REGION Network 5: PODAJANJE PLOŠČICE
   RUNG wire#powerrail
      Contact( #JeVRočnemNačinu )
      { S7_Templates := "SrcType := Int" } EQ_Contact(in1 := #stCilindra, in2 := 5)
      wire#w1
      Contact( #"TIPPEN_-" )
      S_Coil( #"Y1/2" )
      R_Coil( #"Y1/2_2" )
   END_RUNG
   RUNG wire#w1
      Contact( #"TIPPEN_+" )
      Contact( "FB_KEYENCE_GT2_ODMIKVARJENJA".oPoz1Dosezena )
      Contact( "FB_KEYENCE_GT2_ODMIKVARJENJA".oPoz1Dosezena )
      Contact( "Y1/4_odmičniCilinderVarjenje_GOR" )
      R_Coil( #"Y1/2" )
      S_Coil( #"Y1/2_2" )
   END_RUNG
   // the same network as SCL:
   #_w1 := #JeVRočnemNačinu AND (#stCilindra = 5);
   IF #_w1 AND #"TIPPEN_-" THEN
       #"Y1/2" := TRUE;
       #"Y1/2_2" := FALSE;
   END_IF;
   IF #_w1 AND #"TIPPEN_+" AND "FB_KEYENCE_GT2_ODMIKVARJENJA".oPoz1Dosezena AND "FB_KEYENCE_GT2_ODMIKVARJENJA".oPoz1Dosezena AND "Y1/4_odmičniCilinderVarjenje_GOR" THEN
       #"Y1/2" := FALSE;
       #"Y1/2_2" := TRUE;
   END_IF;
END_REGION

REGION Network 6: DVIG/SPUST ELEKTRODE
   RUNG wire#powerrail
      Contact( #JeVRočnemNačinu )
      { S7_Templates := "SrcType := Int" } EQ_Contact(in1 := #stCilindra, in2 := 6)
      wire#w1
      Contact( #"TIPPEN_-" )
      S_Coil( #"Y1/4_1" )
      R_Coil( #"Y1/4_2" )
   END_RUNG
   RUNG wire#w1
      Contact( #"TIPPEN_+" )
      R_Coil( #"Y1/4_1" )
      S_Coil( #"Y1/4_2" )
   END_RUNG
   // the same network as SCL:
   #_w1 := #JeVRočnemNačinu AND (#stCilindra = 6);
   IF #_w1 AND #"TIPPEN_-" THEN
       #"Y1/4_1" := TRUE;
       #"Y1/4_2" := FALSE;
   END_IF;
   IF #_w1 AND #"TIPPEN_+" THEN
       #"Y1/4_1" := FALSE;
       #"Y1/4_2" := TRUE;
   END_IF;
END_REGION

REGION Network 7: PORAVNAVA KONTAKTA
   RUNG wire#powerrail
      Contact( #JeVRočnemNačinu )
      { S7_Templates := "SrcType := Int" } EQ_Contact(in1 := #stCilindra, in2 := 7)
      wire#w1
      Contact( #"TIPPEN_-" )
      S_Coil( #"Y2/3_2" )
      R_Coil( #"Y2/3_1" )
   END_RUNG
   RUNG wire#w1
      Contact( #"TIPPEN_+" )
      R_Coil( #"Y2/3_2" )
      S_Coil( #"Y2/3_1" )
   END_RUNG
   // the same network as SCL:
   #_w1 := #JeVRočnemNačinu AND (#stCilindra = 7);
   IF #_w1 AND #"TIPPEN_-" THEN
       #"Y2/3_2" := TRUE;
       #"Y2/3_1" := FALSE;
   END_IF;
   IF #_w1 AND #"TIPPEN_+" THEN
       #"Y2/3_2" := FALSE;
       #"Y2/3_1" := TRUE;
   END_IF;
END_REGION

REGION Network 8: ODKLEP/ZAKLEP KONUSA - ROTACISKA MIZA
   RUNG wire#powerrail
      Contact( #JeVRočnemNačinu )
      { S7_Templates := "SrcType := Int" } EQ_Contact(in1 := #stCilindra, in2 := 8)
      wire#w1
      Contact( #"TIPPEN_-" )
      R_Coil( #"Y3/1_1" )
   END_RUNG
   RUNG wire#w1
      Contact( #"TIPPEN_+" )
      S_Coil( #"Y3/1_1" )
   END_RUNG
   // the same network as SCL:
   #_w1 := #JeVRočnemNačinu AND (#stCilindra = 8);
   IF #_w1 AND #"TIPPEN_-" THEN #"Y3/1_1" := FALSE; END_IF;
   IF #_w1 AND #"TIPPEN_+" THEN #"Y3/1_1" := TRUE; END_IF;
END_REGION

REGION Network 9: ODKLEP/ZAKLEP VSTAVLJANJA KOMADA V MIZO - ODKLEP ZA VSTAVLJANJE
   RUNG wire#powerrail
      Contact( #JeVRočnemNačinu )
      { S7_Templates := "SrcType := Int" } EQ_Contact(in1 := #stCilindra, in2 := 9)
      wire#w1
      Contact( #"TIPPEN_-" )
      R_Coil( #"Y3/3_1" )
   END_RUNG
   RUNG wire#w1
      Contact( #"TIPPEN_+" )
      S_Coil( #"Y3/3_1" )
   END_RUNG
   // the same network as SCL:
   #_w1 := #JeVRočnemNačinu AND (#stCilindra = 9);
   IF #_w1 AND #"TIPPEN_-" THEN #"Y3/3_1" := FALSE; END_IF;
   IF #_w1 AND #"TIPPEN_+" THEN #"Y3/3_1" := TRUE; END_IF;
END_REGION

REGION Network 10: ODKLEP/ZAKLEP DRŽALA IZMETA KOMADA
   RUNG wire#powerrail
      Contact( #JeVRočnemNačinu )
      { S7_Templates := "SrcType := Int" } EQ_Contact(in1 := #stCilindra, in2 := 10)
      wire#w1
      Contact( #"TIPPEN_-" )
      R_Coil( #"Y4/3_1" )
   END_RUNG
   RUNG wire#w1
      Contact( #"TIPPEN_+" )
      S_Coil( #"Y4/3_1" )
   END_RUNG
   // the same network as SCL:
   #_w1 := #JeVRočnemNačinu AND (#stCilindra = 10);
   IF #_w1 AND #"TIPPEN_-" THEN #"Y4/3_1" := FALSE; END_IF;
   IF #_w1 AND #"TIPPEN_+" THEN #"Y4/3_1" := TRUE; END_IF;
END_REGION

REGION Network 11: IZMET KOMADA
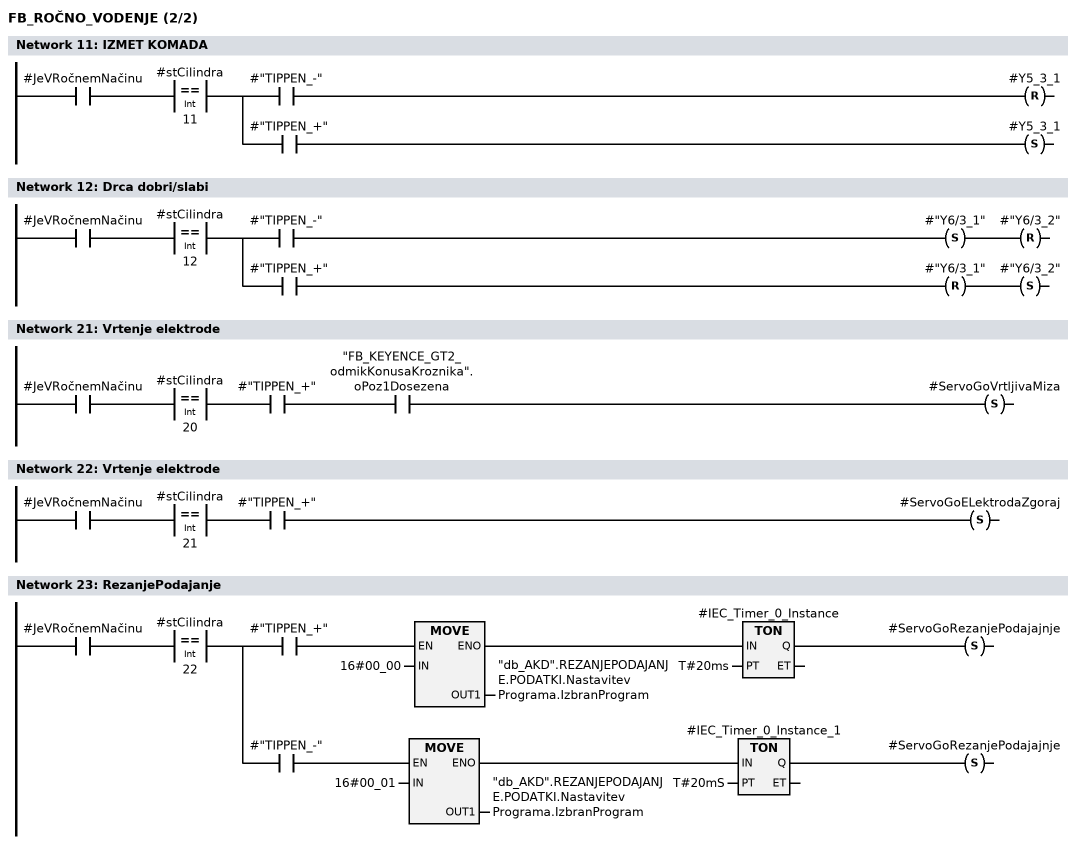
   RUNG wire#powerrail
      Contact( #JeVRočnemNačinu )
      { S7_Templates := "SrcType := Int" } EQ_Contact(in1 := #stCilindra, in2 := 11)
      wire#w1
      Contact( #"TIPPEN_-" )
      R_Coil( #Y5_3_1 )
   END_RUNG
   RUNG wire#w1
      Contact( #"TIPPEN_+" )
      S_Coil( #Y5_3_1 )
   END_RUNG
   // the same network as SCL:
   #_w1 := #JeVRočnemNačinu AND (#stCilindra = 11);
   IF #_w1 AND #"TIPPEN_-" THEN #Y5_3_1 := FALSE; END_IF;
   IF #_w1 AND #"TIPPEN_+" THEN #Y5_3_1 := TRUE; END_IF;
END_REGION

REGION Network 12: Drca dobri/slabi
   RUNG wire#powerrail
      Contact( #JeVRočnemNačinu )
      { S7_Templates := "SrcType := Int" } EQ_Contact(in1 := #stCilindra, in2 := 12)
      wire#w1
      Contact( #"TIPPEN_-" )
      S_Coil( #"Y6/3_1" )
      R_Coil( #"Y6/3_2" )
   END_RUNG
   RUNG wire#w1
      Contact( #"TIPPEN_+" )
      R_Coil( #"Y6/3_1" )
      S_Coil( #"Y6/3_2" )
   END_RUNG
   // the same network as SCL:
   #_w1 := #JeVRočnemNačinu AND (#stCilindra = 12);
   IF #_w1 AND #"TIPPEN_-" THEN
       #"Y6/3_1" := TRUE;
       #"Y6/3_2" := FALSE;
   END_IF;
   IF #_w1 AND #"TIPPEN_+" THEN
       #"Y6/3_1" := FALSE;
       #"Y6/3_2" := TRUE;
   END_IF;
END_REGION

REGION Network 21: Vrtenje elektrode
   RUNG wire#powerrail
      Contact( #JeVRočnemNačinu )
      { S7_Templates := "SrcType := Int" } EQ_Contact(in1 := #stCilindra, in2 := 20)
      Contact( #"TIPPEN_+" )
      Contact( "FB_KEYENCE_GT2_odmikKonusaKroznika".oPoz1Dosezena )
      S_Coil( #ServoGoVrtljivaMiza )
   END_RUNG
   // the same network as SCL:
   IF #JeVRočnemNačinu AND (#stCilindra = 20) AND #"TIPPEN_+" AND "FB_KEYENCE_GT2_odmikKonusaKroznika".oPoz1Dosezena THEN
       #ServoGoVrtljivaMiza := TRUE;
   END_IF;
END_REGION

REGION Network 22: Vrtenje elektrode
   RUNG wire#powerrail
      Contact( #JeVRočnemNačinu )
      { S7_Templates := "SrcType := Int" } EQ_Contact(in1 := #stCilindra, in2 := 21)
      Contact( #"TIPPEN_+" )
      S_Coil( #ServoGoELektrodaZgoraj )
   END_RUNG
   // the same network as SCL:
   IF #JeVRočnemNačinu AND (#stCilindra = 21) AND #"TIPPEN_+" THEN #ServoGoELektrodaZgoraj := TRUE; END_IF;
END_REGION

REGION Network 23: RezanjePodajanje
   #_w1 := #JeVRočnemNačinu AND (#stCilindra = 22);
   #_w2 := #_w1 AND #"TIPPEN_+";
   IF #_w2 THEN "db_AKD".REZANJEPODAJANJE.PODATKI.NastavitevPrograma.IzbranProgram := 16#00_00; END_IF;
   #IEC_Timer_0_Instance(IN := #_w2, PT := T#20ms);   // TON
   IF #IEC_Timer_0_Instance.Q THEN #ServoGoRezanjePodajajnje := TRUE; END_IF;
   #_w3 := #_w1 AND #"TIPPEN_-";
   IF #_w3 THEN "db_AKD".REZANJEPODAJANJE.PODATKI.NastavitevPrograma.IzbranProgram := 16#00_01; END_IF;
   #IEC_Timer_0_Instance_1(IN := #_w3, PT := T#20mS);   // TON
   IF #IEC_Timer_0_Instance_1.Q THEN #ServoGoRezanjePodajajnje := TRUE; END_IF;
END_REGION
END_FUNCTION_BLOCK

FUNCTION_BLOCK "FB_KEYENCE_GT2"   // FB12, LAD
{ S7_Optimized_Access := 'TRUE' }
VERSION : 0.1
   VAR_INPUT
      w_inAddr : DWord;   // VALUE| VALUE|VALUE|BDC1-4
      iPoz1 : DInt;
      iPoz2 : DInt;
      iPoz4 : DInt;
      iPoz3 : DInt;
      HISTEREZA : Int := 800;
      tol1 : Int;
      tol2 : Int;
      tol3 : Int;
      tol4 : Int;
   END_VAR
   VAR_OUTPUT
      out : UDInt;   // Rezultat int
      bBDC1 : Bool;   // Končni položaj 1
      bBDC2 : Bool;   // Končni položaj 2
      bBDC3 : Bool;   // Končni položaj 3
      bBDC4 : Bool;   // Končni položaj 4
      oPoz1Dosezena : Bool;
      oPoz2Dosezena : Bool;
      oPoz3Dosezena : Bool;
      oPoz4Dosezena : Bool;
   END_VAR
   VAR RETAIN
      w_statRor : Word;
      W_ST : Word;
   END_VAR
   VAR
      B0 : Byte;
      B1 : Byte;
   END_VAR
BEGIN

REGION Network 2 (SCL): Rezultat int
   //pozicija dosezena
   //

   #out := #w_inAddr;
   REGION POZICIJA 1
       IF (#iPoz1 - (#HISTEREZA + #tol1)) < #out AND #out < (#iPoz1 + (#HISTEREZA + #tol1)) AND #iPoz1 <> 0 THEN
           #oPoz1Dosezena := true;
   ELSE
       #oPoz1Dosezena := false;
   END_IF;
   END_REGION


   REGION POZICIJA 2
       IF (#iPoz2 - (#HISTEREZA+#tol2)) < #out AND #out < (#iPoz2 + #HISTEREZA+#tol2) AND #iPoz1 <> 0 THEN
       #oPoz2Dosezena := true;
   ELSE
       #oPoz2Dosezena := false;
   END_IF;
   END_REGION

   REGION POZICIJA 3
       IF (#iPoz3 - (#HISTEREZA+#tol3)) < #out AND #out < (#iPoz3 + #HISTEREZA+#tol3) AND #iPoz3 <> 0 THEN
           #oPoz3Dosezena := true;
       ELSE
           #oPoz3Dosezena := false;
       END_IF;
   END_REGION

   REGION POZICIJA 4
       IF (#iPoz4 - (#HISTEREZA+#tol4)) < #out AND #out < (#iPoz4 + #HISTEREZA+#tol4) AND #iPoz4 <> 0 THEN
           #oPoz4Dosezena := true;
       ELSE
           #oPoz4Dosezena := false;
       END_IF;
   END_REGION
END_REGION
END_FUNCTION_BLOCK

FUNCTION_BLOCK "FB_IZMETKOMADA"   // FB13, LAD
{ S7_Optimized_Access := 'TRUE' }
VERSION : 0.1
   VAR_OUTPUT
      VentilZaDržanjeKomada : Bool;
      VentilZaIzmetKomada : Bool;
      DržaDobriSlavi : Bool;
      DržaSlabi : Bool;
   END_VAR
   VAR_IN_OUT
      KomadiPrisotniByte : Byte;
   END_VAR
   VAR RETAIN
      statIzdelekPrisoten : Bool;
      IEC_Timer_0_Instance : TON_TIME;
      IEC_Timer_0_Instance_1 : TON_TIME;
      KoraIzmetaKoncan : Bool;
      merjerji : Array[0..10] of Bool;
   END_VAR
   VAR
      konec : Bool;
   END_VAR
BEGIN

REGION Network 2
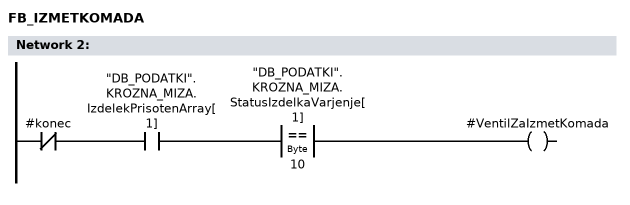
   RUNG wire#powerrail
      I_Contact( #konec )
      Contact( "DB_PODATKI".KROZNA_MIZA.IzdelekPrisotenArray[1] )
      { S7_Templates := "SrcType := Byte" } EQ_Contact(in1 := "DB_PODATKI".KROZNA_MIZA.StatusIzdelkaVarjenje[1], in2 := 10)
      Coil( #VentilZaIzmetKomada )
   END_RUNG
   // the same network as SCL:
   #VentilZaIzmetKomada := NOT #konec AND "DB_PODATKI".KROZNA_MIZA.IzdelekPrisotenArray[1] AND ("DB_PODATKI".KROZNA_MIZA.StatusIzdelkaVarjenje[1] = 10);
END_REGION
END_FUNCTION_BLOCK

FUNCTION_BLOCK "FB_VstavljanjeIzdelkaVMizo"   // FB14, LAD
{ S7_Optimized_Access := 'TRUE' }
VERSION : 0.1
   VAR_INPUT
      PogojZaVstavljanje : Bool;   // Ko na mizi ni komada
   END_VAR
   VAR_OUTPUT
      IzdelekVstavljenVMizo : Bool;
   END_VAR
   VAR RETAIN
      Korak : UInt;
   END_VAR
   VAR
      Ton : Array[0..1] of TON_TIME;
   END_VAR
   VAR_TEMP   // added for the SCL form of the ladder/FBD networks
      _w1 : Bool;
   END_VAR
BEGIN

REGION Network 1: ČajanjeZaVstavljanje
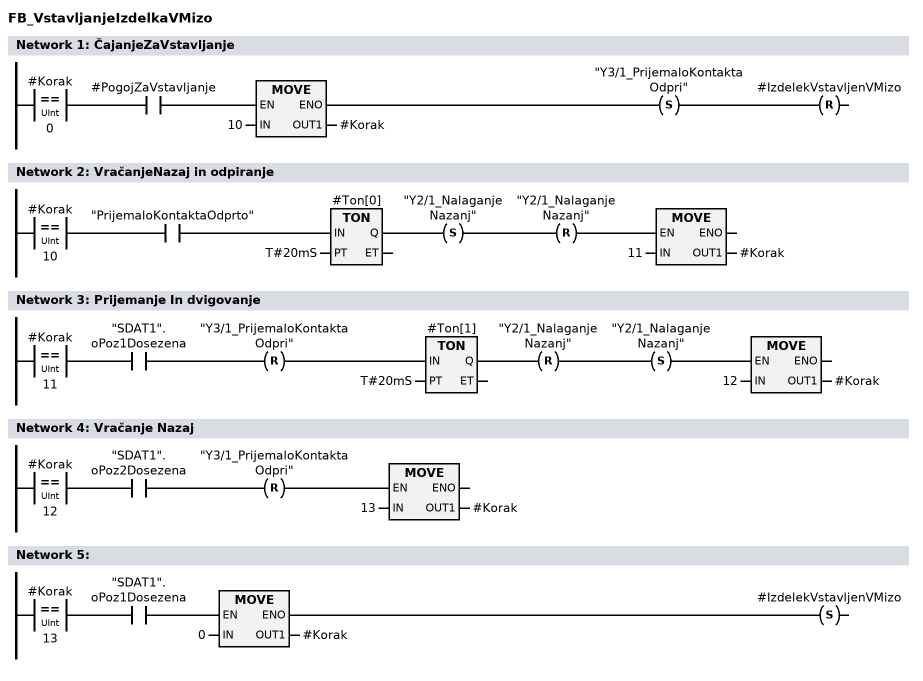
   RUNG wire#powerrail
      { S7_Templates := "SrcType := UInt" } EQ_Contact(in1 := #Korak, in2 := 0)
      Contact( #PogojZaVstavljanje )
      Move(in := 10, out1 => #Korak)
      S_Coil( "Y3/1_PrijemaloKontaktaOdpri" )
      R_Coil( #IzdelekVstavljenVMizo )
   END_RUNG
   // the same network as SCL:
   #_w1 := (#Korak = 0) AND #PogojZaVstavljanje;
   IF #_w1 THEN
       #Korak := 10;
       "Y3/1_PrijemaloKontaktaOdpri" := TRUE;
       #IzdelekVstavljenVMizo := FALSE;
   END_IF;
END_REGION

REGION Network 2: VračanjeNazaj in odpiranje
   #Ton[0].TON(IN := (#Korak = 10) AND "PrijemaloKontaktaOdprto", PT := T#20mS);
   IF #Ton[0].Q THEN
       "Y2/1_NalaganjeNazanj" := TRUE;
       "Y2/1_NalaganjeNazanj" := FALSE;
       #Korak := 11;
   END_IF;
END_REGION

REGION Network 3: Prijemanje In dvigovanje
   #_w1 := (#Korak = 11) AND "SDAT1".oPoz1Dosezena;
   IF #_w1 THEN "Y3/1_PrijemaloKontaktaOdpri" := FALSE; END_IF;
   #Ton[1].TON(IN := #_w1, PT := T#20mS);
   IF #Ton[1].Q THEN
       "Y2/1_NalaganjeNazanj" := FALSE;
       "Y2/1_NalaganjeNazanj" := TRUE;
       #Korak := 12;
   END_IF;
END_REGION

REGION Network 4: Vračanje Nazaj
   RUNG wire#powerrail
      { S7_Templates := "SrcType := UInt" } EQ_Contact(in1 := #Korak, in2 := 12)
      Contact( "SDAT1".oPoz2Dosezena )
      R_Coil( "Y3/1_PrijemaloKontaktaOdpri" )
      Move(in := 13, out1 => #Korak)
   END_RUNG
   // the same network as SCL:
   IF (#Korak = 12) AND "SDAT1".oPoz2Dosezena THEN
       "Y3/1_PrijemaloKontaktaOdpri" := FALSE;
       #Korak := 13;
   END_IF;
END_REGION

REGION Network 5
   RUNG wire#powerrail
      { S7_Templates := "SrcType := UInt" } EQ_Contact(in1 := #Korak, in2 := 13)
      Contact( "SDAT1".oPoz1Dosezena )
      Move(in := 0, out1 => #Korak)
      S_Coil( #IzdelekVstavljenVMizo )
   END_RUNG
   // the same network as SCL:
   #_w1 := (#Korak = 13) AND "SDAT1".oPoz1Dosezena;
   IF #_w1 THEN
       #Korak := 0;
       #IzdelekVstavljenVMizo := TRUE;
   END_IF;
END_REGION
END_FUNCTION_BLOCK

FUNCTION_BLOCK "FB_IOL_BANNER"   // FB15, LAD
{ S7_Optimized_Access := 'TRUE' }
VERSION : 0.1
   VAR_INPUT
      Color1 : Byte;
      ColorFlashRate : Byte;
      Color2 : Byte;
      AudioMode : Byte;
      Rotation : Bool;
      ANimationType : Byte;
      Color1Intensity : Byte;
      Color2Intensety : Byte;
   END_VAR
   VAR_OUTPUT
      oWord : DWord;
      oByte0 : Byte;
      oByte1 : Byte;
      oByte2 : Byte;
      oByte3 : Byte;
   END_VAR
   VAR
      bytes : Array[0..3] of Byte;
   END_VAR
BEGIN

REGION Network 2 (SCL)
   #bytes[0] := #Color1 + SHL(IN := #ColorFlashRate, N := 5);
   #bytes[1] := #Color2 + SHL(IN := #AudioMode, N := 5);
   #bytes[2] := #ANimationType + SHL(IN := #Color1Intensity, N := 4);
   #bytes[3] := #Color2Intensety;
   //#oWord :=#bytes[0]+SHL(IN:=#bytes[1],N:=8);
   //#oWord := ROL(IN := #oWord, N := 0);

   #oByte0 := #bytes[0];
   #oByte1 := #bytes[1];
   #oByte2 := #bytes[2];
   #oByte3 := #bytes[3];
END_REGION
END_FUNCTION_BLOCK

FUNCTION_BLOCK "FB_TekociTrak"   // FB16, LAD
{ S7_Optimized_Access := 'TRUE' }
VERSION : 0.1
   VAR_INPUT
      i_StetjeKosov : Bool;
      i_ON_OFF_TekociTrak : Bool;
      i_stevecSlabihKosov : UInt;
      i_MAX_SKATLA1 : UInt;
      i_MAX_SKATLA2 : UInt;
      i_IzprazniSKatlo1 : Bool;
      i_iprazniSkatlo2 : Bool;
   END_VAR
   VAR_OUTPUT
      o_TekočiTrak : Bool;
      o_PolnjenjeSkatle2 : Bool;
      o_Skatla1Polna : Bool;
      o_Skatla2Polna : Bool;
   END_VAR
   VAR_IN_OUT
      i_StevecSkatle1 : UInt;
      i_StevecSkatle2 : UInt;
      i_ResetNapake : Bool;
   END_VAR
   VAR RETAIN
      stat_skatla1Polna : Bool;
      stat_skatla2Polna : Bool;
      merkerji : Array[0..3] of Bool;
      IEC_Timer_0_Instance : TON_TIME;
      IEC_Timer_0_Instance_1 : TON_TIME;
      SkatliPolni : Bool;
      statPolnjenjeSkatle2 : Bool;
   END_VAR
   VAR_TEMP   // added for the SCL form of the ladder/FBD networks
      _w1 : Bool;
      _w2 : Bool;
      _w3 : Bool;
      _w4 : Bool;
   END_VAR
BEGIN

REGION Network 1: Vklop Tekocega Traka
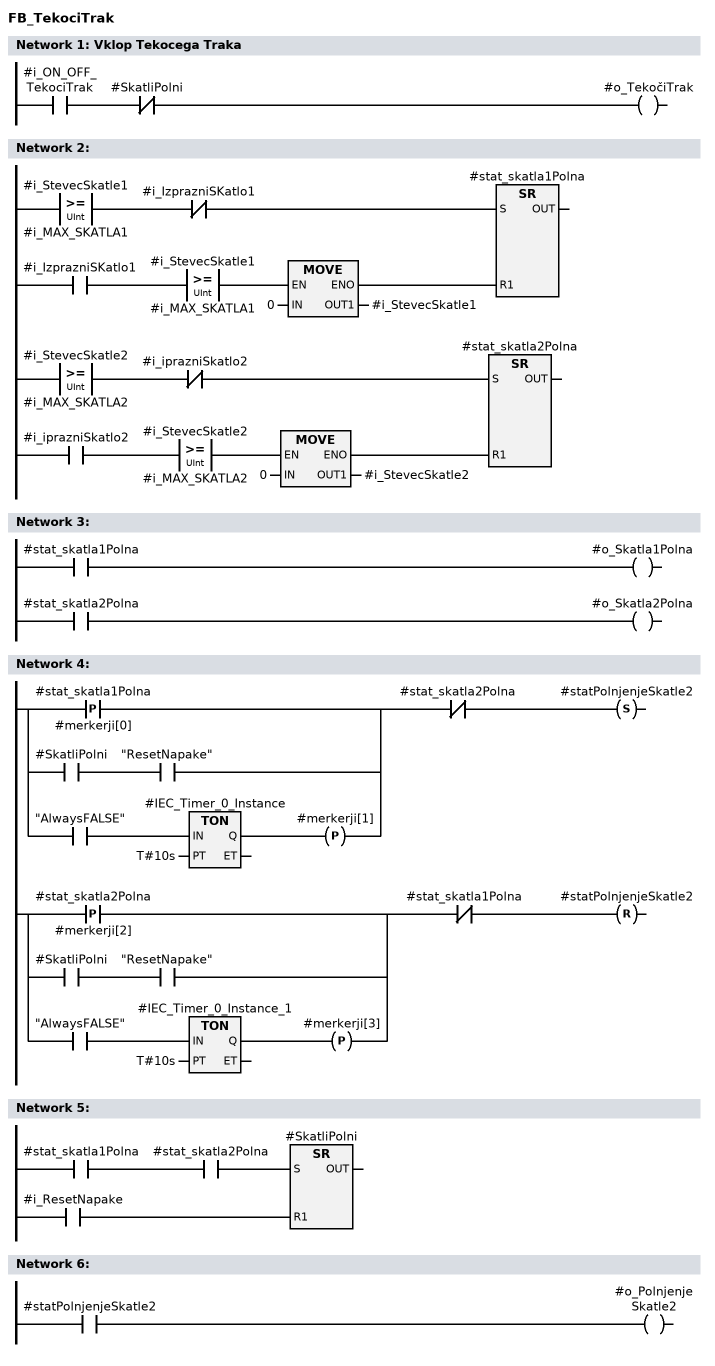
   RUNG wire#powerrail
      Contact( #i_ON_OFF_TekociTrak )
      I_Contact( #SkatliPolni )
      Coil( #o_TekočiTrak )
   END_RUNG
   // the same network as SCL:
   #o_TekočiTrak := #i_ON_OFF_TekociTrak AND NOT #SkatliPolni;
END_REGION

REGION Network 2
   RUNG wire#powerrail
      { S7_Templates := "SrcType := UInt" } GE_Contact(in1 := #i_StevecSkatle1, in2 := #i_MAX_SKATLA1)
      I_Contact( #i_IzprazniSKatlo1 )
      S_SR(operand := #stat_skatla1Polna, r1 := wire#w1)
   END_RUNG
   RUNG wire#powerrail
      Contact( #i_IzprazniSKatlo1 )
      { S7_Templates := "SrcType := UInt" } GE_Contact(in1 := #i_StevecSkatle1, in2 := #i_MAX_SKATLA1)
      Move(in := 0, out1 => #i_StevecSkatle1)
   END_RUNG wire#w1
   RUNG wire#powerrail
      { S7_Templates := "SrcType := UInt" } GE_Contact(in1 := #i_StevecSkatle2, in2 := #i_MAX_SKATLA2)
      I_Contact( #i_iprazniSkatlo2 )
      S_SR(operand := #stat_skatla2Polna, r1 := wire#w2)
   END_RUNG
   RUNG wire#powerrail
      Contact( #i_iprazniSkatlo2 )
      { S7_Templates := "SrcType := UInt" } GE_Contact(in1 := #i_StevecSkatle2, in2 := #i_MAX_SKATLA2)
      Move(in := 0, out1 => #i_StevecSkatle2)
   END_RUNG wire#w2
   // the same network as SCL:
   #_w1 := #i_IzprazniSKatlo1 AND (#i_StevecSkatle1 >= #i_MAX_SKATLA1);
   #_w2 := (#i_StevecSkatle1 >= #i_MAX_SKATLA1) AND NOT #i_IzprazniSKatlo1;
   IF #_w1 THEN #i_StevecSkatle1 := 0; END_IF;
   IF #_w2 THEN
       #stat_skatla1Polna := TRUE;   // SR flip-flop
   END_IF;
   IF #_w1 THEN #stat_skatla1Polna := FALSE; END_IF;
   #_w3 := #i_iprazniSkatlo2 AND (#i_StevecSkatle2 >= #i_MAX_SKATLA2);
   #_w4 := (#i_StevecSkatle2 >= #i_MAX_SKATLA2) AND NOT #i_iprazniSkatlo2;
   IF #_w3 THEN #i_StevecSkatle2 := 0; END_IF;
   IF #_w4 THEN
       #stat_skatla2Polna := TRUE;   // SR flip-flop
   END_IF;
   IF #_w3 THEN #stat_skatla2Polna := FALSE; END_IF;
END_REGION

REGION Network 3
   RUNG wire#powerrail
      Contact( #stat_skatla1Polna )
      Coil( #o_Skatla1Polna )
   END_RUNG
   RUNG wire#powerrail
      Contact( #stat_skatla2Polna )
      Coil( #o_Skatla2Polna )
   END_RUNG
   // the same network as SCL:
   #o_Skatla1Polna := #stat_skatla1Polna;
   #o_Skatla2Polna := #stat_skatla2Polna;
END_REGION

REGION Network 4
   #_w1 := #stat_skatla1Polna AND NOT #merkerji[0];   // rising edge of #stat_skatla1Polna
   #merkerji[0] := #stat_skatla1Polna;
   #IEC_Timer_0_Instance(IN := "AlwaysFALSE", PT := T#10s);   // TON
   #_w2 := #IEC_Timer_0_Instance.Q AND NOT #merkerji[1];   // rising edge
   #merkerji[1] := #IEC_Timer_0_Instance.Q;
   IF (#_w1 OR (#SkatliPolni AND "ResetNapake") OR #_w2) AND NOT #stat_skatla2Polna THEN
       #statPolnjenjeSkatle2 := TRUE;
   END_IF;
   #_w3 := #stat_skatla2Polna AND NOT #merkerji[2];   // rising edge of #stat_skatla2Polna
   #merkerji[2] := #stat_skatla2Polna;
   #IEC_Timer_0_Instance_1(IN := "AlwaysFALSE", PT := T#10s);   // TON
   #_w4 := #IEC_Timer_0_Instance_1.Q AND NOT #merkerji[3];   // rising edge
   #merkerji[3] := #IEC_Timer_0_Instance_1.Q;
   IF (#_w3 OR (#SkatliPolni AND "ResetNapake") OR #_w4) AND NOT #stat_skatla1Polna THEN
       #statPolnjenjeSkatle2 := FALSE;
   END_IF;
END_REGION

REGION Network 5
   RUNG wire#powerrail
      Contact( #stat_skatla1Polna )
      Contact( #stat_skatla2Polna )
      S_SR(operand := #SkatliPolni, r1 := wire#w1)
   END_RUNG
   RUNG wire#powerrail
      Contact( #i_ResetNapake )
   END_RUNG wire#w1
   // the same network as SCL:
   IF #stat_skatla1Polna AND #stat_skatla2Polna THEN
       #SkatliPolni := TRUE;   // SR flip-flop
   END_IF;
   IF #i_ResetNapake THEN #SkatliPolni := FALSE; END_IF;
END_REGION

REGION Network 6
   RUNG wire#powerrail
      Contact( #statPolnjenjeSkatle2 )
      Coil( #o_PolnjenjeSkatle2 )
   END_RUNG
   // the same network as SCL:
   #o_PolnjenjeSkatle2 := #statPolnjenjeSkatle2;
END_REGION
END_FUNCTION_BLOCK

FUNCTION_BLOCK "FB_TIMERS"   // FB17, LAD
{ S7_Optimized_Access := 'TRUE' }
VERSION : 0.1
   VAR_INPUT
      TriggerCycleTime : Bool;
   END_VAR
   VAR RETAIN
      IEC_Timer_0_Instance : TONR_TIME;
      merkerji : Array[0..1] of Bool;
      TimerOn : Bool;
   END_VAR
   VAR
      timerarray : Array[0..1] of LDT;
      IEC_Timer_0_Instance_1 : TON_TIME;
      "WORD" : Word;
   END_VAR
   VAR RETAIN
      "counter" : Int;
   END_VAR
   VAR
      "TIME" : LDT;
      cycleTime : LTime;
      counterstevca : DInt;
      one : Bool;
      CycleTimeTIe : Time;
      TImeint : Int;
      TimeReal : Real;
      TIME_1 : Real;
      mm : Int;
   END_VAR
   VAR RETAIN
      IzdelkiNaUro : Int;
   END_VAR
   VAR
      staticmm : Int;
      realmm : Real;
      intfloor : Int;
   END_VAR
   VAR_TEMP
      IZRACUNAJ : Bool;
      SUB : Real;
      "MOD" : Real;
      nn : LReal;
   END_VAR
   VAR_TEMP   // added for the SCL form of the ladder/FBD networks
      _w1 : Bool;
      _w2 : Bool;
      _w3 : Bool;
   END_VAR
BEGIN

REGION Network 1
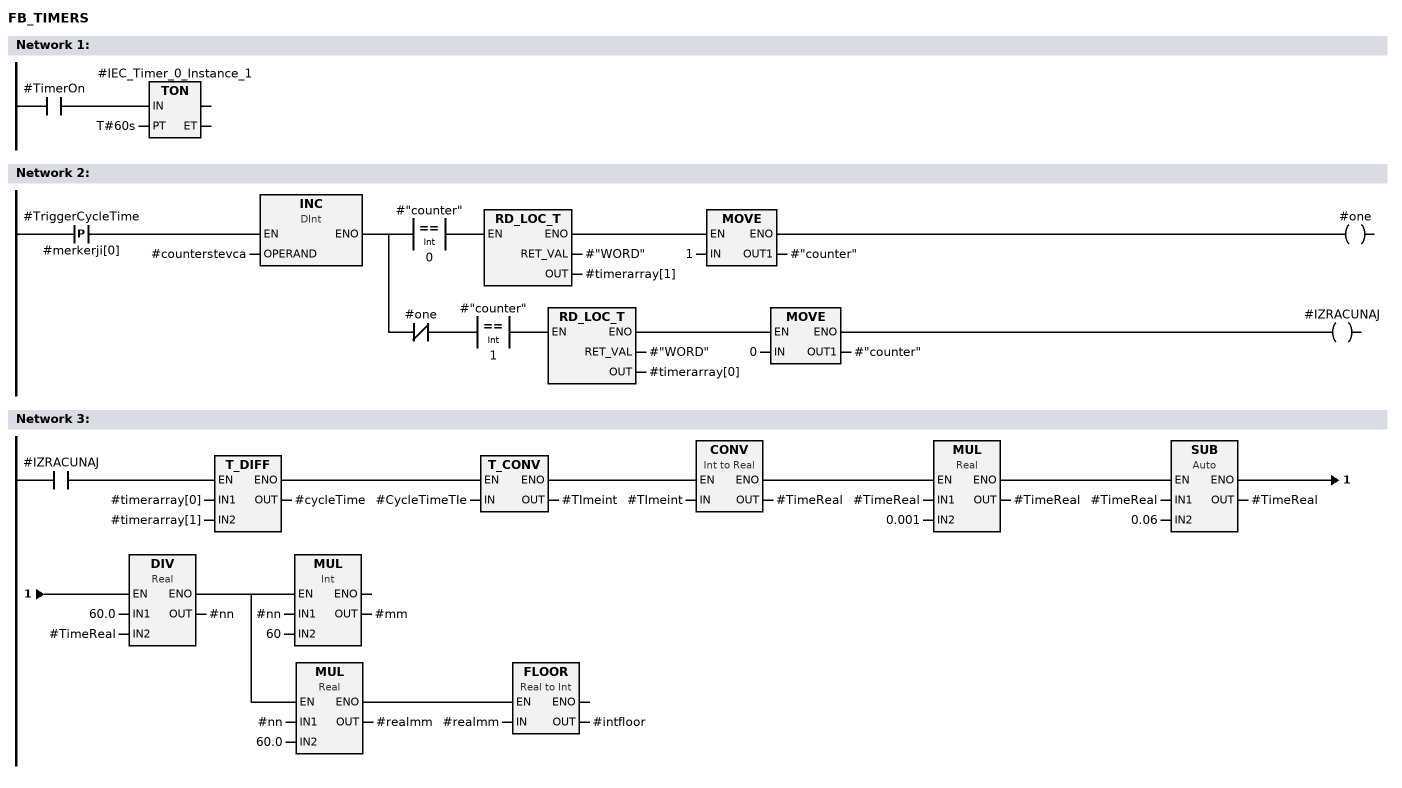
   #IEC_Timer_0_Instance_1(IN := #TimerOn, PT := T#60s);   // TON
END_REGION

REGION Network 2
   // ENO of a box is taken as its EN; it also drops when the box reports an error
   #_w1 := #TriggerCycleTime AND NOT #merkerji[0];   // rising edge of #TriggerCycleTime
   #merkerji[0] := #TriggerCycleTime;
   IF #_w1 THEN #counterstevca := #counterstevca + 1; END_IF;
   #_w2 := #_w1 AND (#"counter" = 0);
   IF #_w2 THEN
       #"WORD" := RD_LOC_T(OUT => #timerarray[1]);
       #"counter" := 1;
   END_IF;
   #one := #_w2;
   #_w3 := #_w1 AND NOT #one AND (#"counter" = 1);
   IF #_w3 THEN
       #"WORD" := RD_LOC_T(OUT => #timerarray[0]);
       #"counter" := 0;
   END_IF;
   #IZRACUNAJ := #_w3;
END_REGION

REGION Network 3
   // ENO of a box is taken as its EN; it also drops when the box reports an error
   IF #IZRACUNAJ THEN
       #cycleTime := T_DIFF(IN1 := #timerarray[0], IN2 := #timerarray[1]);
       #TImeint := T_CONV(IN := #CycleTimeTIe);
       #TimeReal := INT_TO_REAL(#TImeint);
       #TimeReal := #TimeReal * 0.001;
       #TimeReal := #TimeReal - 0.06;
       #nn := 60.0 / #TimeReal;
       #mm := #nn * 60;
       #realmm := #nn * 60.0;
       #intfloor := FLOOR(#realmm);
   END_IF;
END_REGION

REGION Network 5 (SCL)
   #CycleTimeTIe := LTIME_TO_TIME(IN := #cycleTime);
   #staticmm := #mm;
END_REGION
END_FUNCTION_BLOCK

FUNCTION_BLOCK "Block_1"   // FB18, ProDiag
{ S7_Optimized_Access := 'TRUE' }
VERSION : 0.1
   VAR
      PC_Flags : PC_Flags_V2;
      State : SV_FB_State_V2;
      "FB_GL_PROGRAM_DB.#Vstavljanje v mizo.VA_Merr_1" : SV_State_V2;
      "Type_Mess_E_C1_1052700-2064" : Diag_Alarm_2;
      "FB_GL_PROGRAM_DB.#Vstavljanje v mizo_1.VA_Merr_1" : SV_State_V2;
      "FB_GL_PROGRAM_DB.#Step40.VA_Merr_1" : SV_State_V2;
      "FB_GL_PROGRAM_DB.#PODAJANJE PLOŠČICE.VA_Mtxt_1" : SV_State_V2;
      "Type_Mess_T_C1_1052700-2064" : Diag_Alarm_2;
   END_VAR
   VAR_TEMP
      t_TempSvStateUDT : SV_State_V2;
      t_TempAlarmInstance : <type 200004f>;
      t_TempAsocValue1 : Variant;
      t_TempAsocValue2 : Variant;
      t_TempAsocValue3 : Variant;
   END_VAR
BEGIN
END_FUNCTION_BLOCK

FUNCTION_BLOCK "FB_LocalTime"   // FB19, LAD
{ S7_Optimized_Access := 'TRUE' }
VERSION : 0.1
   VAR_INPUT
      bWriteLocalTime : Bool;
   END_VAR
   VAR
      DateAndTIME : LDT;
      RD_LOC_T_err : Word;
      WR_LOC : Struct
         LOCALTIME : LDT;
         DST : Bool;
         ret_val : Word;
      END_STRUCT;
   END_VAR
BEGIN

REGION Network 1
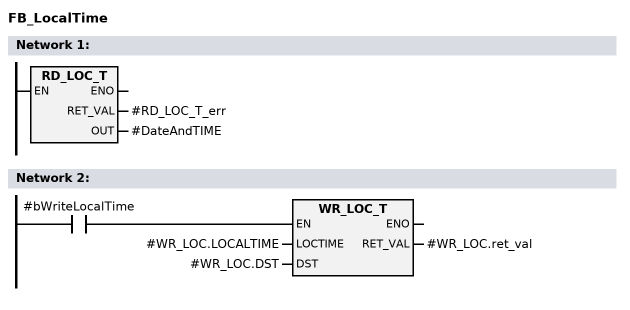
   #RD_LOC_T_err := RD_LOC_T(OUT => #DateAndTIME);
END_REGION

REGION Network 2
   IF #bWriteLocalTime THEN
       #WR_LOC.ret_val := WR_LOC_T(LOCTIME := #WR_LOC.LOCALTIME, DST := #WR_LOC.DST);
   END_IF;
END_REGION
END_FUNCTION_BLOCK

FUNCTION_BLOCK "FB_KAMERA_TRIG"   // FB20, LAD
{ S7_Optimized_Access := 'TRUE' }
VERSION : 0.1
   VAR_INPUT
      bCameraTrig : Bool;   // Pogoj za kamera triger
      bCameraFeedback : Bool;   // Kamera OK/NOK - feedback iz kamere
   END_VAR
   VAR_OUTPUT
      Out1Trig : Bool;   // Triger za izhod kamera
      Out2Trig : Bool;   // Triger za izhod kamere
   END_VAR
   VAR_IN_OUT
      io_StatusArrayCamere : Byte;   // Krožna miza - status kamere
   END_VAR
   VAR RETAIN
      stat_CamLastValue : Bool;   // kamera zadnji status
      trig : Array[0..1] of Bool;
      korak : Int;
      StatCamArray : Array[0..7] of Bool;
   END_VAR
   VAR_TEMP   // added for the SCL form of the ladder/FBD networks
      _w1 : Bool;
   END_VAR
BEGIN

REGION Network 1: Triger kamere 500mS
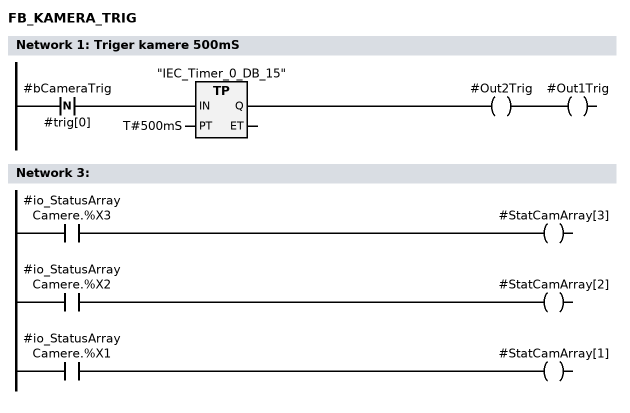
   #_w1 := NOT #bCameraTrig AND #trig[0];   // falling edge of #bCameraTrig
   #trig[0] := #bCameraTrig;
   "IEC_Timer_0_DB_15".TP(IN := #_w1, PT := T#500mS);
   #Out2Trig := "IEC_Timer_0_DB_15".Q;
   #Out1Trig := "IEC_Timer_0_DB_15".Q;
END_REGION

REGION Network 2 (SCL): 0 - NOK, 1 OK
   "F_TRIG_DB_CAMERATRIG"(CLK:=#bCameraTrig);

   IF "F_TRIG_DB_CAMERATRIG".Q THEN //negativni triger
       //ČE STA vrednosti različni postavi izhod na "1" - kamera je OK - kamera naredi toggle, če je izhod OK
       IF #stat_CamLastValue XOR #bCameraFeedback THEN
           #io_StatusArrayCamere.%X3:= 1;
       ELSE
           #io_StatusArrayCamere.%X3 := 0;
       END_IF;
       //shranjevanje zadnje vrednosti
       #stat_CamLastValue := #bCameraFeedback; 
   END_IF;
END_REGION

REGION Network 3
   RUNG wire#powerrail
      Contact( #io_StatusArrayCamere.%X3 )
      Coil( #StatCamArray[3] )
   END_RUNG
   RUNG wire#powerrail
      Contact( #io_StatusArrayCamere.%X2 )
      Coil( #StatCamArray[2] )
   END_RUNG
   RUNG wire#powerrail
      Contact( #io_StatusArrayCamere.%X1 )
      Coil( #StatCamArray[1] )
   END_RUNG
   // the same network as SCL:
   #StatCamArray[3] := #io_StatusArrayCamere.%X3;
   #StatCamArray[2] := #io_StatusArrayCamere.%X2;
   #StatCamArray[1] := #io_StatusArrayCamere.%X1;
END_REGION
END_FUNCTION_BLOCK

FUNCTION "FC_SHIFTREGISTRI" : Void   // FC1, LAD
{ S7_Optimized_Access := 'TRUE' }
VERSION : 0.1
   VAR_INPUT
      TrigerMizaZavrtena : Bool;
      TrigerZavarjeno : Bool;
      ZavarjenoOK : Bool;
      bIzdelekVstavljenVMizo : Bool;   // Izdelek je vstavljen postavi bit na 1
      bTrigIzmetKomada : Bool;
   END_VAR
   VAR_IN_OUT
      IzdelekPrisotenVMizi : Byte;
      IzdelekZavarjen : Byte;
      IzdelekKameraOk : Byte;
      ioStatusIzdelka : Array[0..7] of Byte;
   END_VAR
   VAR_TEMP   // added for the SCL form of the ladder/FBD networks
      _w1 : Bool;
      _w2 : Bool;
   END_VAR
BEGIN

REGION Network 1
   // 1 - nalozeno
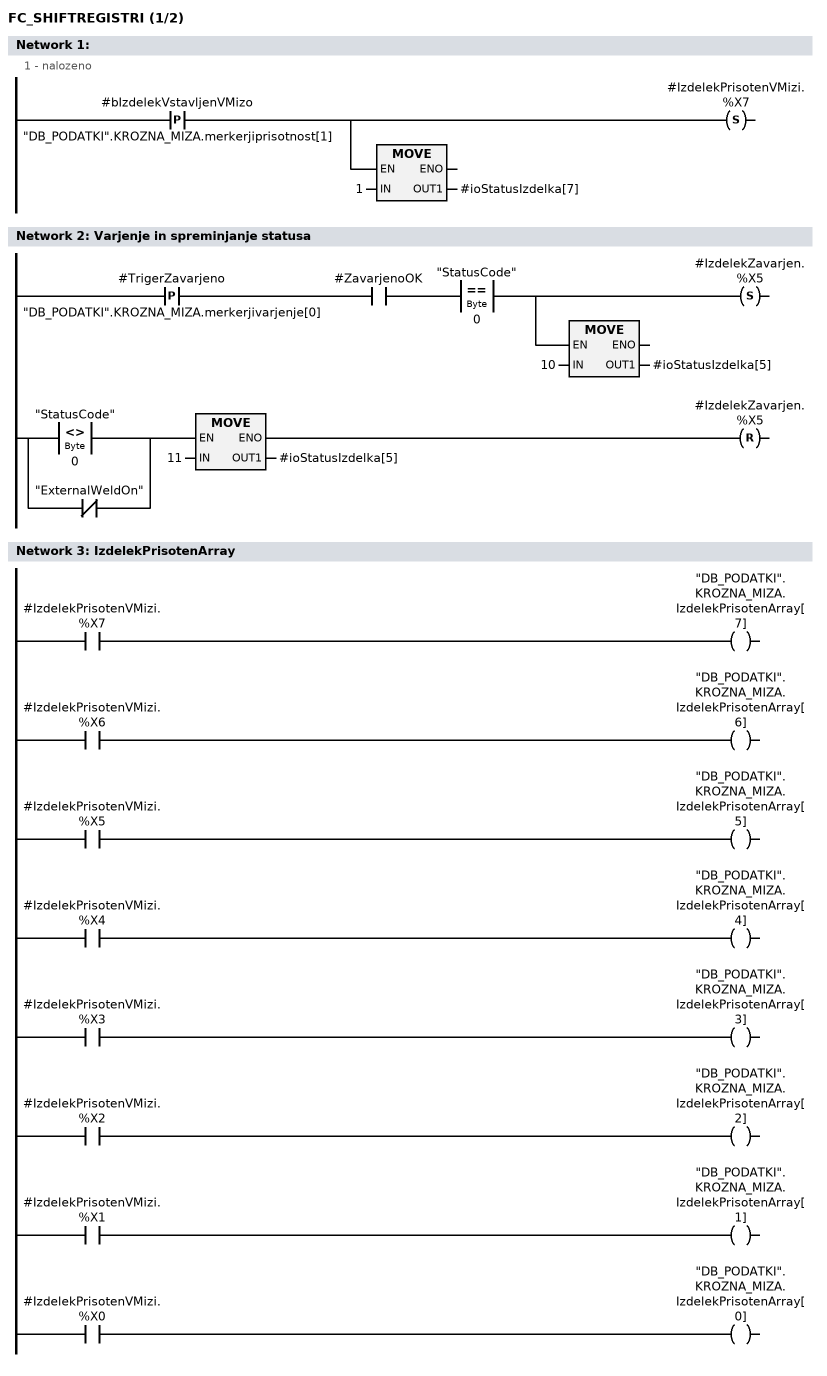
   RUNG wire#powerrail
      P_Contact(operand := #bIzdelekVstavljenVMizo, bit := "DB_PODATKI".KROZNA_MIZA.merkerjiprisotnost[1])
      wire#w1
      S_Coil( #IzdelekPrisotenVMizi.%X7 )
   END_RUNG
   RUNG wire#w1
      Move(in := 1, out1 => #ioStatusIzdelka[7])
   END_RUNG
   // the same network as SCL:
   #_w1 := #bIzdelekVstavljenVMizo AND NOT "DB_PODATKI".KROZNA_MIZA.merkerjiprisotnost[1];   // rising edge of #bIzdelekVstavljenVMizo
   "DB_PODATKI".KROZNA_MIZA.merkerjiprisotnost[1] := #bIzdelekVstavljenVMizo;
   IF #_w1 THEN
       #IzdelekPrisotenVMizi.%X7 := TRUE;
       #ioStatusIzdelka[7] := 1;
   END_IF;
END_REGION

REGION Network 2: Varjenje in spreminjanje statusa
   RUNG wire#powerrail
      P_Contact(operand := #TrigerZavarjeno, bit := "DB_PODATKI".KROZNA_MIZA.merkerjivarjenje[0])
      Contact( #ZavarjenoOK )
      { S7_Templates := "SrcType := Byte" } EQ_Contact(in1 := "StatusCode", in2 := 0)
      wire#w1
      S_Coil( #IzdelekZavarjen.%X5 )
   END_RUNG
   RUNG wire#w1
      Move(in := 10, out1 => #ioStatusIzdelka[5])
   END_RUNG
   RUNG wire#powerrail
      { S7_Templates := "SrcType := Byte" } NE_Contact(in1 := "StatusCode", in2 := 0)
      wire#w2
      Move(in := 11, out1 => #ioStatusIzdelka[5])
      R_Coil( #IzdelekZavarjen.%X5 )
   END_RUNG
   RUNG wire#powerrail
      I_Contact( "ExternalWeldOn" )
   END_RUNG wire#w2
   // the same network as SCL:
   #_w1 := #TrigerZavarjeno AND NOT "DB_PODATKI".KROZNA_MIZA.merkerjivarjenje[0];   // rising edge of #TrigerZavarjeno
   "DB_PODATKI".KROZNA_MIZA.merkerjivarjenje[0] := #TrigerZavarjeno;
   IF #_w1 AND #ZavarjenoOK AND ("StatusCode" = 0) THEN
       #IzdelekZavarjen.%X5 := TRUE;
       #ioStatusIzdelka[5] := 10;
   END_IF;
   IF ("StatusCode" <> 0) OR NOT "ExternalWeldOn" THEN
       #ioStatusIzdelka[5] := 11;
       #IzdelekZavarjen.%X5 := FALSE;
   END_IF;
END_REGION

REGION Network 3: IzdelekPrisotenArray
   RUNG wire#powerrail
      Contact( #IzdelekPrisotenVMizi.%X7 )
      Coil( "DB_PODATKI".KROZNA_MIZA.IzdelekPrisotenArray[7] )
   END_RUNG
   RUNG wire#powerrail
      Contact( #IzdelekPrisotenVMizi.%X6 )
      Coil( "DB_PODATKI".KROZNA_MIZA.IzdelekPrisotenArray[6] )
   END_RUNG
   RUNG wire#powerrail
      Contact( #IzdelekPrisotenVMizi.%X5 )
      Coil( "DB_PODATKI".KROZNA_MIZA.IzdelekPrisotenArray[5] )
   END_RUNG
   RUNG wire#powerrail
      Contact( #IzdelekPrisotenVMizi.%X4 )
      Coil( "DB_PODATKI".KROZNA_MIZA.IzdelekPrisotenArray[4] )
   END_RUNG
   RUNG wire#powerrail
      Contact( #IzdelekPrisotenVMizi.%X3 )
      Coil( "DB_PODATKI".KROZNA_MIZA.IzdelekPrisotenArray[3] )
   END_RUNG
   RUNG wire#powerrail
      Contact( #IzdelekPrisotenVMizi.%X2 )
      Coil( "DB_PODATKI".KROZNA_MIZA.IzdelekPrisotenArray[2] )
   END_RUNG
   RUNG wire#powerrail
      Contact( #IzdelekPrisotenVMizi.%X1 )
      Coil( "DB_PODATKI".KROZNA_MIZA.IzdelekPrisotenArray[1] )
   END_RUNG
   RUNG wire#powerrail
      Contact( #IzdelekPrisotenVMizi.%X0 )
      Coil( "DB_PODATKI".KROZNA_MIZA.IzdelekPrisotenArray[0] )
   END_RUNG
   // the same network as SCL:
   "DB_PODATKI".KROZNA_MIZA.IzdelekPrisotenArray[7] := #IzdelekPrisotenVMizi.%X7;
   "DB_PODATKI".KROZNA_MIZA.IzdelekPrisotenArray[6] := #IzdelekPrisotenVMizi.%X6;
   "DB_PODATKI".KROZNA_MIZA.IzdelekPrisotenArray[5] := #IzdelekPrisotenVMizi.%X5;
   "DB_PODATKI".KROZNA_MIZA.IzdelekPrisotenArray[4] := #IzdelekPrisotenVMizi.%X4;
   "DB_PODATKI".KROZNA_MIZA.IzdelekPrisotenArray[3] := #IzdelekPrisotenVMizi.%X3;
   "DB_PODATKI".KROZNA_MIZA.IzdelekPrisotenArray[2] := #IzdelekPrisotenVMizi.%X2;
   "DB_PODATKI".KROZNA_MIZA.IzdelekPrisotenArray[1] := #IzdelekPrisotenVMizi.%X1;
   "DB_PODATKI".KROZNA_MIZA.IzdelekPrisotenArray[0] := #IzdelekPrisotenVMizi.%X0;
END_REGION

REGION Network 5
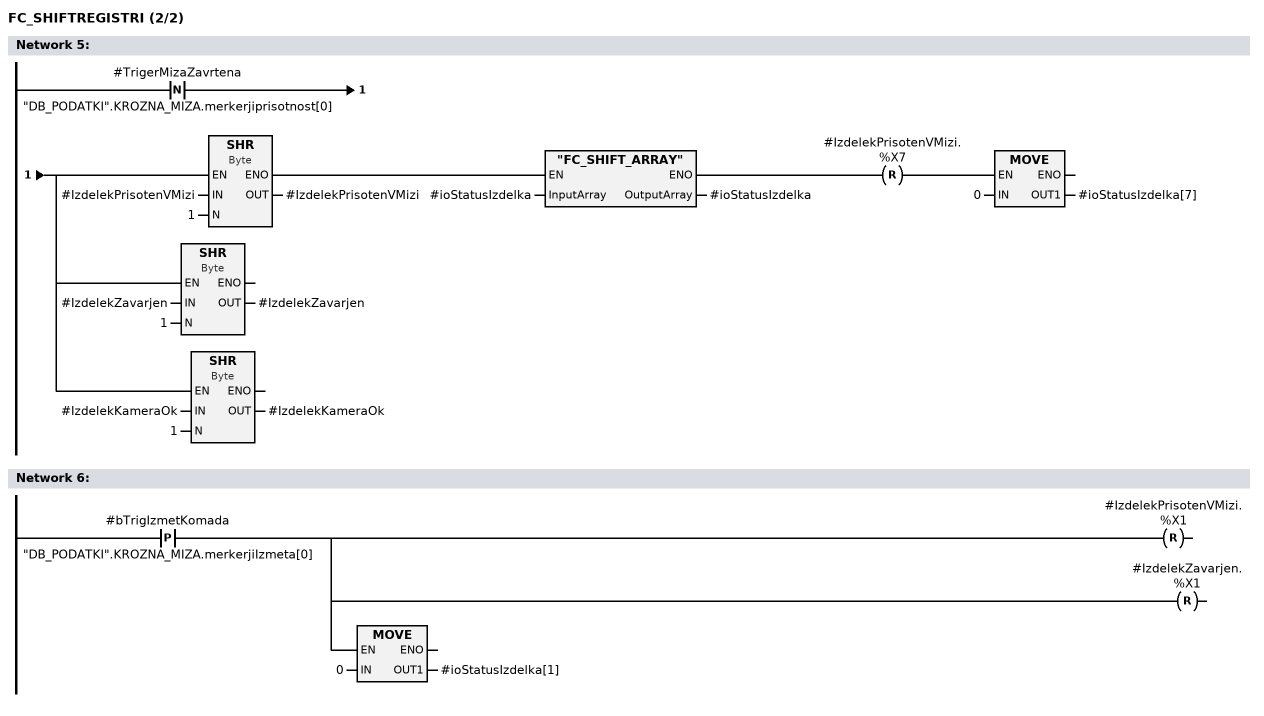
   RUNG wire#powerrail
      N_Contact(operand := #TrigerMizaZavrtena, bit := "DB_PODATKI".KROZNA_MIZA.merkerjiprisotnost[0])
      wire#w1
      { S7_Templates := "SrcType := Byte" } Shr(in := #IzdelekPrisotenVMizi, n := 1, out => #IzdelekPrisotenVMizi)
      "FC_SHIFT_ARRAY"(InputArray := #ioStatusIzdelka, OutputArray => #ioStatusIzdelka)
      R_Coil( #IzdelekPrisotenVMizi.%X7 )
      Move(in := 0, out1 => #ioStatusIzdelka[7])
   END_RUNG
   RUNG wire#w1
      { S7_Templates := "SrcType := Byte" } Shr(in := #IzdelekZavarjen, n := 1, out => #IzdelekZavarjen)
   END_RUNG
   RUNG wire#w1
      { S7_Templates := "SrcType := Byte" } Shr(in := #IzdelekKameraOk, n := 1, out => #IzdelekKameraOk)
   END_RUNG
   // the same network as SCL:
   #_w1 := NOT #TrigerMizaZavrtena AND "DB_PODATKI".KROZNA_MIZA.merkerjiprisotnost[0];   // falling edge of #TrigerMizaZavrtena
   "DB_PODATKI".KROZNA_MIZA.merkerjiprisotnost[0] := #TrigerMizaZavrtena;
   IF #_w1 THEN #IzdelekPrisotenVMizi := SHR(IN := #IzdelekPrisotenVMizi, N := 1); END_IF;
   "FC_SHIFT_ARRAY"(EN := #_w1, InputArray := #ioStatusIzdelka, OutputArray => #ioStatusIzdelka, ENO => #_w2);
   IF #_w2 THEN
       #IzdelekPrisotenVMizi.%X7 := FALSE;
       #ioStatusIzdelka[7] := 0;
   END_IF;
   IF #_w1 THEN
       #IzdelekZavarjen := SHR(IN := #IzdelekZavarjen, N := 1);
       #IzdelekKameraOk := SHR(IN := #IzdelekKameraOk, N := 1);
   END_IF;
END_REGION

REGION Network 6
   RUNG wire#powerrail
      P_Contact(operand := #bTrigIzmetKomada, bit := "DB_PODATKI".KROZNA_MIZA.merkerjiIzmeta[0])
      wire#w1
      R_Coil( #IzdelekPrisotenVMizi.%X1 )
   END_RUNG
   RUNG wire#w1
      R_Coil( #IzdelekZavarjen.%X1 )
   END_RUNG
   RUNG wire#w1
      Move(in := 0, out1 => #ioStatusIzdelka[1])
   END_RUNG
   // the same network as SCL:
   #_w1 := #bTrigIzmetKomada AND NOT "DB_PODATKI".KROZNA_MIZA.merkerjiIzmeta[0];   // rising edge of #bTrigIzmetKomada
   "DB_PODATKI".KROZNA_MIZA.merkerjiIzmeta[0] := #bTrigIzmetKomada;
   IF #_w1 THEN
       #IzdelekPrisotenVMizi.%X1 := FALSE;
       #IzdelekZavarjen.%X1 := FALSE;
       #ioStatusIzdelka[1] := 0;
   END_IF;
END_REGION
END_FUNCTION

FUNCTION "FC_VARJENJE" : Void   // FC2, LAD
{ S7_Optimized_Access := 'TRUE' }
VERSION : 0.1
   VAR_INPUT
      ZahtevaZaVarjenje : Bool;
      IzbiraProgram : Byte;
      VarilniTokOn : Bool;   // 0 OFF | 1 ON
      VarjenjePogoji : Bool;
      iVarjenjeKončano : Bool;
      VklopSpotSelection : Bool;
      i_bResetWithWC : Bool;
      i_bResetWithReweld : Bool;
   END_VAR
   VAR_OUTPUT
      VarjenjeGO : Bool;
      Program : Byte;
      oVarilniTokOn : Bool;
      oSpotSelection : Bool;
      o_bResetWithWC : Bool;
      o_bResetWithReweld : Bool;
   END_VAR
BEGIN

REGION Network 1: Vklop varjenja
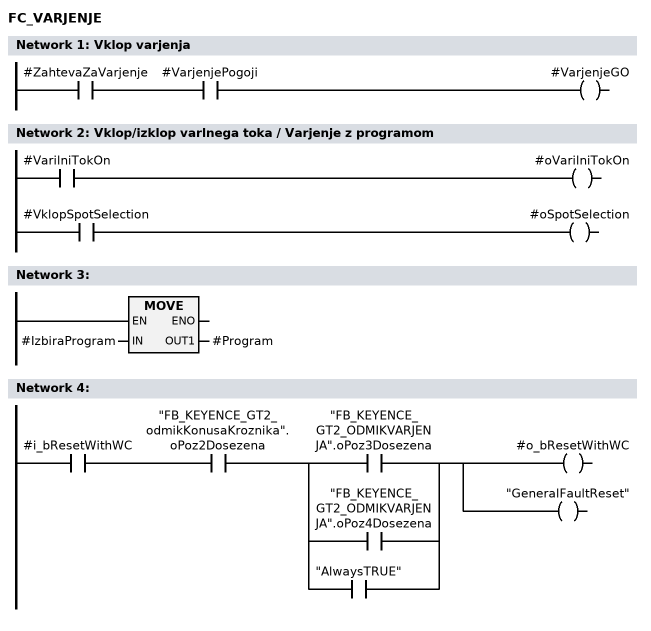
   RUNG wire#powerrail
      Contact( #ZahtevaZaVarjenje )
      Contact( #VarjenjePogoji )
      Coil( #VarjenjeGO )
   END_RUNG
   // the same network as SCL:
   #VarjenjeGO := #ZahtevaZaVarjenje AND #VarjenjePogoji;
END_REGION

REGION Network 2: Vklop/izklop varlnega toka / Varjenje z programom
   RUNG wire#powerrail
      Contact( #VarilniTokOn )
      Coil( #oVarilniTokOn )
   END_RUNG
   RUNG wire#powerrail
      Contact( #VklopSpotSelection )
      Coil( #oSpotSelection )
   END_RUNG
   // the same network as SCL:
   #oVarilniTokOn := #VarilniTokOn;
   #oSpotSelection := #VklopSpotSelection;
END_REGION

REGION Network 3
   RUNG wire#powerrail
      Move(in := #IzbiraProgram, out1 => #Program)
   END_RUNG
   // the same network as SCL:
   #Program := #IzbiraProgram;
END_REGION

REGION Network 4
   RUNG wire#powerrail
      Contact( #i_bResetWithWC )
      Contact( "FB_KEYENCE_GT2_odmikKonusaKroznika".oPoz2Dosezena )
      wire#w1
      Contact( "FB_KEYENCE_GT2_ODMIKVARJENJA".oPoz3Dosezena )
      wire#w2
      Coil( #o_bResetWithWC )
   END_RUNG
   RUNG wire#w1
      Contact( "FB_KEYENCE_GT2_ODMIKVARJENJA".oPoz4Dosezena )
   END_RUNG wire#w2
   RUNG wire#w1
      Contact( "AlwaysTRUE" )
   END_RUNG wire#w2
   RUNG wire#w2
      Coil( "GeneralFaultReset" )
   END_RUNG
   // the same network as SCL:
   #o_bResetWithWC := #i_bResetWithWC AND "FB_KEYENCE_GT2_odmikKonusaKroznika".oPoz2Dosezena AND ("FB_KEYENCE_GT2_ODMIKVARJENJA".oPoz3Dosezena OR "FB_KEYENCE_GT2_ODMIKVARJENJA".oPoz4Dosezena OR "AlwaysTRUE");
   "GeneralFaultReset" := #o_bResetWithWC;
END_REGION
END_FUNCTION

FUNCTION "FC_BTN_INDIKACIJA" : Void   // FC3, LAD
{ S7_Optimized_Access := 'TRUE' }
VERSION : 0.1
   VAR_INPUT
      inError : Bool;
      inAutomaticMode : Bool;
      RUN : Bool;
      iPogojiZaRun : Bool;
   END_VAR
   VAR_OUTPUT
      ErrorLed : Bool;
      RunLed : Bool;
   END_VAR
BEGIN

